text list "Banner_ManIntMsg2": 0 '**Local Message Display**'; 1 '~Spare MB2[0].1'; 2 '~Spare MB2[0].2'; 3 '~Spare MB2[0].3'; 4 '~Spare MB2[0].4'; 5 '~Spare MB2[0].5'; 6 '~Spare MB2[0].6'; 7 '~Spare MB2[0].7'; 8 '~Spare MB2[0].8'; 9 '~Spare MB2[0].9'; 10 '~Spare MB2[0].10'; 11 '~Spare MB2[0].11'; 12 '~Spare MB2[0].12'; 13 '~Spare MB2[0].13'; 14 '~Spare MB2[0].14'; 15 '~Spare MB2[0].15'; 16 '~Spare MB2[0].16'; 17 '~Spare MB2[0].17'; 18 '~Spare MB2[0].18'; 19 '~Spare MB2[0].19'; 20 '~Spare MB2[0].20'; 21 '~Spare MB2[0].21'; 22 '~Spare MB2[0].22'; 23 '~Spare MB2[0].23'; 24 '~Spare MB2[0].24'; 25 '~Spare MB2[0].25'; 26 '~Spare MB2[0].26'; 27 '~Spare MB2[0].27'; 28 '~Spare MB2[0].28'; 29 '~Spare MB2[0].29'; 30 '~Spare MB2[0].30'; 31 '~Spare MB2[0].31'; 32 '~PDPES1 - PDP EtherNet Switch Connection Inhibited MB2[1].0'; 33 '~Spare MB2[1].1'; 34 '~Spare MB2[1].2'; 35 '~MPES1 - Main Panel EtherNet Switch Connection Inhibited MB2[1].3'; 36 '~Spare MB2[1].4'; 37 '~Spare MB2[1].5'; 38 '~MPES2 - Main Panel EtherNet Switch Connection Inhibited MB2[1].6'; 39 '~Spare MB2[1].7'; 40 '~Spare MB2[1].8'; 41 '~MPES3 - Main Panel EtherNet Switch Connection Inhibited MB2[1].9'; 42 '~Spare MB2[1].10'; 43 '~Spare MB2[1].11'; 44 '~Spare MB2[1].12'; 45 '~Spare MB2[1].13'; 46 '~Spare MB2[1].14'; 47 '~Spare MB2[1].15'; 48 '~Spare MB2[1].16'; 49 '~MPES1 - Main Panel Control Power Disconnect Not On MB2[1].17'; 50 '~PDP 1 - Panel Output Disconnect Safety Switch Not On MB2[1].18'; 51 '~PDP 2 - Panel Output Disconnect Safety Switch Not On MB2[1].19'; 52 '~PDP 3 - Panel Output Disconnect Safety Switch Not On MB2[1].20'; 53 '~Spare MB2[1].21'; 54 '~Spare MB2[1].22'; 55 '~Spare MB2[1].23'; 56 '~Spare MB2[1].24'; 57 '~Spare MB2[1].25'; 58 '~Spare MB2[1].26'; 59 '~Spare MB2[1].27'; 60 '~Spare MB2[1].28'; 61 '~Spare MB2[1].29'; 62 '~Spare MB2[1].30'; 63 '~Spare MB2[1].31'; 64 '~ES3ES1 - ES3 EtherNet Switch Connection Inhibited MB2[2].0'; 65 '~Spare MB2[2].1'; 66 '~Spare MB2[2].2'; 67 '~Spare MB2[2].3'; 68 '~Spare MB2[2].4'; 69 '~Spare MB2[2].5'; 70 '~Spare MB2[2].6'; 71 '~Spare MB2[2].7'; 72 '~Spare MB2[2].8'; 73 '~ES3Sfty - Motion Control Enable Relay #1 MECR1 Still On MB2[2].9'; 74 '~ES3Sfty - Motion Control Enable Relay #1 MECR1 Not On MB2[2].10'; 75 '~ES3Sfty - Motion Control Enable Relay #2 MECR2 Still On MB2[2].11'; 76 '~ES3Sfty - Motion Control Enable Relay #2 MECR2 Not On MB2[2].12'; 77 '~ES3Sfty - EtherNet Switch Sfty Relays RESSR1 RESSR2 Not On MB2[2].13'; 78 '~ES3Sfty - EtherNet Switch Sfty Relays RESSR1 RESSR2 Still On MB2[2].14'; 79 '~Spare MB2[2].15'; 80 '~Spare MB2[2].16'; 81 '~Spare MB2[2].17'; 82 '~Spare MB2[2].18'; 83 '~Spare MB2[2].19'; 84 '~ES3 S003 Safety Gate #1 Open MB2[2].20'; 85 '~ES3 S003 Safety Gate #2 Open MB2[2].21'; 86 '~Spare MB2[2].22'; 87 '~Spare MB2[2].23'; 88 '~Spare MB2[2].24'; 89 '~Spare MB2[2].25'; 90 '~Spare MB2[2].26'; 91 '~Spare MB2[2].27'; 92 '~Spare MB2[2].28'; 93 '~Spare MB2[2].29'; 94 '~Spare MB2[2].30'; 95 '~Spare MB2[2].31'; 96 '~ES4ES1 - ES4 EtherNet Switch Connection Inhibited MB2[3].0'; 97 '~Spare MB2[3].1'; 98 '~Spare MB2[3].2'; 99 '~Spare MB2[3].3'; 100 '~Spare MB2[3].4'; 101 '~Spare MB2[3].5'; 102 '~Spare MB2[3].6'; 103 '~Spare MB2[3].7'; 104 '~Spare MB2[3].8'; 105 '~ES2Sfty - Motion Control Enable Relay #1 MECR1 Still On MB2[3].9'; 106 '~ES2Sfty - Motion Control Enable Relay #1 MECR1 Not On MB2[3].10'; 107 '~ES2Sfty - Motion Control Enable Relay #2 MECR2 Still On MB2[3].11'; 108 '~ES2Sfty - Motion Control Enable Relay #2 MECR2 Not On MB2[3].12'; 109 '~ES2Sfty - EtherNet Switch Sfty Relays RESSR1 RESSR2 Not On MB2[3].13'; 110 '~ES2Sfty - EtherNet Switch Sfty Relays RESSR1 RESSR2 Still On MB2[3].14'; 111 '~Spare MB2[3].15'; 112 '~Spare MB2[3].16'; 113 '~Spare MB2[3].17'; 114 '~Spare MB2[3].18'; 115 '~Spare MB2[3].19'; 116 '~ES2 S002 Safety Gate #1 Open MB2[3].20'; 117 '~ES2 S002 Safety Gate #2 Open MB2[3].21'; 118 '~Spare MB2[3].22'; 119 '~Spare MB2[3].23'; 120 '~Spare MB2[3].24'; 121 '~Spare MB2[3].25'; 122 '~Spare MB2[3].26'; 123 '~Spare MB2[3].27'; 124 '~Spare MB2[3].28'; 125 '~Spare MB2[3].29'; 126 '~Spare MB2[3].30'; 127 '~Spare MB2[3].31'; 128 '~PV3ES1 - PV3 EtherNet Switch Connection Inhibited MB2[4].0'; 129 '~Spare MB2[4].1'; 130 '~Spare MB2[4].2'; 131 '~Spare MB2[4].3'; 132 '~Spare MB2[4].4'; 133 '~Spare MB2[4].5'; 134 '~Spare MB2[4].6'; 135 '~Spare MB2[4].7'; 136 '~Spare MB2[4].8'; 137 '~Spare MB2[4].9'; 138 '~Spare MB2[4].10'; 139 '~PV1Sfty - EtherNet Switch Sfty Relays RESSR1 RESSR2 Not On MB2[4].11'; 140 '~PV1Sfty - EtherNet Switch Sfty Relays RESSR1 RESSR2 Still On MB2[4].12'; 141 '~Spare MB2[4].13'; 142 '~Spare MB2[4].14'; 143 '~PV1 S002 E-Stop Depressed MB2[4].15'; 144 '~PV1 S002 Safety Gate #1 Open MB2[4].16'; 145 '~PV1 S002 Safety Gate #2 Open MB2[4].17'; 146 '~Spare MB2[4].18'; 147 '~Spare MB2[4].19'; 148 '~Spare MB2[4].20'; 149 '~Spare MB2[4].21'; 150 '~Spare MB2[4].22'; 151 '~Spare MB2[4].23'; 152 '~S002 Both PanelViews Have Manual Selected MB2[4].24'; 153 '~S002 PanelView 1 Manual Selected MB2[4].25'; 154 '~Spare MB2[4].26'; 155 '~Spare MB2[4].27'; 156 '~PV1 S002 Auto Not Selected MB2[4].28'; 157 '~PV1 S002 Not In Auto Or Manual MB2[4].29'; 158 '~Spare MB2[4].30'; 159 '~Spare MB2[4].31'; 160 '~PV4ES1 - PV4 EtherNet Switch Connection Inhibited MB2[5].0'; 161 '~Spare MB2[5].1'; 162 '~Spare MB2[5].2'; 163 '~Spare MB2[5].3'; 164 '~Spare MB2[5].4'; 165 '~Spare MB2[5].5'; 166 '~Spare MB2[5].6'; 167 '~Spare MB2[5].7'; 168 '~Spare MB2[5].8'; 169 '~Spare MB2[5].9'; 170 '~Spare MB2[5].10'; 171 '~PV2Sfty - EtherNet Switch Sfty Relays RESSR1 RESSR2 Not On MB2[5].11'; 172 '~PV2Sfty - EtherNet Switch Sfty Relays RESSR1 RESSR2 Still On MB2[5].12'; 173 '~Spare MB2[5].13'; 174 '~Spare MB2[5].14'; 175 '~PV2 S002 PanelView E-Stop Depressed MB2[5].15'; 176 '~PV2 S002 Safety Gate #1 Open MB2[5].16'; 177 '~PV2 S002 Safety Gate #2 Open MB2[5].17'; 178 '~Spare MB2[5].18'; 179 '~Spare MB2[5].19'; 180 '~Spare MB2[5].20'; 181 '~Spare MB2[5].21'; 182 '~Spare MB2[5].22'; 183 '~Spare MB2[5].23'; 184 '~Spare MB2[5].24'; 185 '~S002 PanelView 2 Manual Selected MB2[5].25'; 186 '~Spare MB2[5].26'; 187 '~Spare MB2[5].27'; 188 '~PV2 S002 Auto Not Selected MB2[5].28'; 189 '~PV2 S002 Not In Auto Or Manual MB2[5].29'; 190 '~Spare MB2[5].30'; 191 '~Spare MB2[5].31'; 192 '~S001R09ES1 - S001R09 EtherNet Switch Connection Inhibited MB2[6].0'; 193 '~Spare MB2[6].1'; 194 '~Spare MB2[6].2'; 195 '~Spare MB2[6].3'; 196 '~Spare MB2[6].4'; 197 '~Spare MB2[6].5'; 198 '~Spare MB2[6].6'; 199 '~Spare MB2[6].7'; 200 '~Spare MB2[6].8'; 201 '~Spare MB2[6].9'; 202 '~Spare MB2[6].10'; 203 '~Spare MB2[6].11'; 204 '~Spare MB2[6].12'; 205 '~Spare MB2[6].13'; 206 '~Spare MB2[6].14'; 207 '~Spare MB2[6].15'; 208 '~Spare MB2[6].16'; 209 '~S001R09Sfty - Robot E-Stop Depressed MB2[6].17'; 210 '~S001R09Sfty - Robot Safety Interface Not Enabled MB2[6].18'; 211 '~S001R09Sfty - Robot DCS Has Been Edited MB2[6].19'; 212 '~S001R09CN - Robot Controller Connection Inhibited MB2[6].20'; 213 '~S001R09E#B# - Robot End Effector Module Connection Inhibited MB2[6].21'; 214 '~S001R09E#B# - Robot End Effector Module Connection Inhibited MB2[6].22'; 215 '~S001R09E#B# - Robot End Effector Module Connection Inhibited MB2[6].23'; 216 '~S001R09E#B# - Robot End Effector Module Connection Inhibited MB2[6].24'; 217 '~S001R09E#B# - Robot End Effector Module Connection Inhibited MB2[6].25'; 218 '~S001R09E#B# - Robot End Effector Module Connection Inhibited MB2[6].26'; 219 '~S001R09E#B# - Robot End Effector Module Connection Inhibited MB2[6].27'; 220 '~S001R09E#B# - Robot End Effector Module Connection Inhibited MB2[6].28'; 221 '~S001R09E#B# - Robot End Effector Module Connection Inhibited MB2[6].29'; 222 '~Spare MB2[6].30'; 223 '~Spare MB2[6].31'; 224 '~Spare MB2[7].0'; 225 '~S001R09F#B# - Robot Process I/O Connection Inhibited MB2[7].1'; 226 '~S001R09F#B# - Robot Process I/O Connection Inhibited MB2[7].2'; 227 '~S001R09F#B# - Robot Process I/O Connection Inhibited MB2[7].3'; 228 '~S001R09F#B# - Robot Process I/O Connection Inhibited MB2[7].4'; 229 '~Spare MB2[7].5'; 230 '~Spare MB2[7].6'; 231 '~Spare MB2[7].7'; 232 '~Spare MB2[7].8'; 233 '~Spare MB2[7].9'; 234 '~S001R09CN.I.Safety - Chain Fault MB2[7].10'; 235 '~S001R09CN.I.AirOn - Robot Air Not On MB2[7].11'; 236 '~S001R09CN.I.RbtAuto - Robot Not in Auto MB2[7].12'; 237 '~S001R09CN.M.InTeach - Robot In Teach MB2[7].13'; 238 '~S001R09CN.I.AtMaintPos - Robot At Maintenace MB2[7].14'; 239 '~S001R09CN.I.RunEnblInterruptAck - Robot In Hold MB2[7].15'; 240 '~S001R09CN.M.MaintPosSeld - Robot Maintenance Selected MB2[7].16'; 241 '~Spare MB2[7].17'; 242 '~Spare MB2[7].18'; 243 '~Spare MB2[7].19'; 244 '~S001R09CN.I.ExtAppCommFlt - Robot Application Communication Fault MB2[7].20'; 245 '~S001R09CN.M.AbortPickupSeld - Robot Abort Pickup Selected MB2[7].21'; 246 '~S001R09CN.M.RetFmPounceSeld - Robot Return From Pounce Selected MB2[7].22'; 247 '~S001R09CN.I.StudWld1 Comm Not OK MB2[7].23'; 248 '~S001R09CN.I.StudWld2 Comm Not OK MB2[7].24'; 249 '~S001R09CN.I.WldMode - Robot In No Weld MB2[7].25'; 250 '~S001R09CN.I.PulledTipBypSS - Robot Pulled Tip Bypass Selected MB2[7].26'; 251 '~S001R09CN.I.FlowNoFlowSS - Robot In No Flow MB2[7].27'; 252 '~S001R09CN.I.RvtNoRvtSS - Robot In No Rivet MB2[7].28'; 253 '~S001R09CN.I.WldCtrlCommOk1 - Robot Weld Controller 1 Comm Not OK MB2[7].29'; 254 '~S001R09CN.I.WldModeStud - Robot In No Weld Stud MB2[7].30'; 255 '~S001R09CN.Ix.MigWldNoWld - Robot In No Weld Mig MB2[7].31'; 256 '~S001R09CN.I.StudWld1Rdy - Robot Stud Weld Controller 1 Not Ready MB2[8].0'; 257 '~S001R09CN.I.Rvt1RdyToOperate - Robot Rivet Controller 1 Not Ready MB2[8].1'; 258 '~S001R09CN.Ix.MigRdy - Robot Mig Weld Controller Not Ready MB2[8].2'; 259 '~S001R09CN.Ix.MigWldNoWld - Robot In No Weld MB2[8].3'; 260 '~Spare MB2[8].4'; 261 '~S001R09CN.I.WldCtrlCommOk2 - Robot Weld Controller 2 Comm Not OK MB2[8].5'; 262 '~Spare MB2[8].6'; 263 '~Spare MB2[8].7'; 264 '~S001R09CN.I.StudWld2Rdy - Robot Stud Weld Controller 2 Not Ready MB2[8].8'; 265 '~S001R09CN.I.Rvt2RdyToOperate - Robot Rivet Controller 2 Not Ready MB2[8].9'; 266 '~S001R09CN.Ix.LaserWldOn - Robot Laser In No Cut MB2[8].10'; 267 '~S001R09CN.Ix.GlassNotPres - Robot Laser Glass Not Present MB2[8].11'; 268 '~S001R09CN.Ix.LaserHeadRdy - Robot Laser Head Not Ready MB2[8].12'; 269 '~S001R09CN.Ix.ChillerOn - Robot Laser Chiller Not On MB2[8].13'; 270 '~S001R09CN.Ix.GasOn - Robot Gas Not On MB2[8].14'; 271 '~S001R09 Power Meter Not Ready MB2[8].15'; 272 '~S001R09 No Wire Present Replace Barrel MB2[8].16'; 273 '~S001R09 Wire Feeder Fault Timer MB2[8].17'; 274 '~S001R09CN.Ix.NRFlt - Robot Nut Runner Not Ready MB2[8].18'; 275 '~Spare MB2[8].19'; 276 '~S001R09CN.M.WrongRivetAtNose - Remove Wrong Rivet At Nose MB2[8].20'; 277 '~S001R09CN.M.DisableRbtDrvs - In Rivet Zone But Riveter Not In Auto MB2[8].21'; 278 '~S001R09CN.I.Rvt1SystemInAuto - Rivet Controller 1 Not In Auto MB2[8].22'; 279 '~S001R09CN.I.Rvt2SystemInAuto - Rivet Controller 2 Not In Auto MB2[8].23'; 280 '~S001R09CN.M.RvtC1ReelCtr.DN - Reel Change Required MB2[8].24'; 281 '~S001R09CN.M.RvtC2ReelCtr.DN - Reel Change Required MB2[8].25'; 282 '~S001R09CN.M.AbortSkipRemain - SkipRemaining Aborted, Reset At Rbt Controller Is Required MB2[8].26'; 283 '~Spare MB2[8].27'; 284 '~Spare MB2[8].28'; 285 '~Spare MB2[8].29'; 286 '~Spare MB2[8].30'; 287 '~Spare MB2[8].31'; 288 '~Spare MB2[9].0'; 289 '~Spare MB2[9].1'; 290 '~Spare MB2[9].2'; 291 '~Spare MB2[9].3'; 292 '~Spare MB2[9].4'; 293 '~Spare MB2[9].5'; 294 '~Spare MB2[9].6'; 295 '~Spare MB2[9].7'; 296 '~Spare MB2[9].8'; 297 '~Spare MB2[9].9'; 298 '~Spare MB2[9].10'; 299 '~Spare MB2[9].11'; 300 '~Spare MB2[9].12'; 301 '~Spare MB2[9].13'; 302 '~Spare MB2[9].14'; 303 '~Spare MB2[9].15'; 304 '~Spare MB2[9].16'; 305 '~Spare MB2[9].17'; 306 '~Spare MB2[9].18'; 307 '~Spare MB2[9].19'; 308 '~Spare MB2[9].20'; 309 '~Spare MB2[9].21'; 310 '~Spare MB2[9].22'; 311 '~Spare MB2[9].23'; 312 '~Spare MB2[9].24'; 313 '~Spare MB2[9].25'; 314 '~Spare MB2[9].26'; 315 '~Spare MB2[9].27'; 316 '~Spare MB2[9].28'; 317 '~Spare MB2[9].29'; 318 '~Spare MB2[9].30'; 319 '~Spare MB2[9].31'; 320 '~Spare MB2[10].0'; 321 '~Spare MB2[10].1'; 322 '~Spare MB2[10].2'; 323 '~Spare MB2[10].3'; 324 '~Spare MB2[10].4'; 325 '~Spare MB2[10].5'; 326 '~Spare MB2[10].6'; 327 '~Spare MB2[10].7'; 328 '~Spare MB2[10].8'; 329 '~Spare MB2[10].9'; 330 '~Spare MB2[10].10'; 331 '~Spare MB2[10].11'; 332 '~Spare MB2[10].12'; 333 '~Spare MB2[10].13'; 334 '~Spare MB2[10].14'; 335 '~Spare MB2[10].15'; 336 '~Spare MB2[10].16'; 337 '~Spare MB2[10].17'; 338 '~Spare MB2[10].18'; 339 '~Spare MB2[10].19'; 340 '~Spare MB2[10].20'; 341 '~Spare MB2[10].21'; 342 '~Spare MB2[10].22'; 343 '~Spare MB2[10].23'; 344 '~Spare MB2[10].24'; 345 '~Spare MB2[10].25'; 346 '~Spare MB2[10].26'; 347 '~Spare MB2[10].27'; 348 '~Spare MB2[10].28'; 349 '~Spare MB2[10].29'; 350 '~Spare MB2[10].30'; 351 '~Spare MB2[10].31'; 352 '~Spare MB2[11].0'; 353 '~Spare MB2[11].1'; 354 '~Spare MB2[11].2'; 355 '~Spare MB2[11].3'; 356 '~Spare MB2[11].4'; 357 '~Spare MB2[11].5'; 358 '~Spare MB2[11].6'; 359 '~Spare MB2[11].7'; 360 '~Spare MB2[11].8'; 361 '~Spare MB2[11].9'; 362 '~Spare MB2[11].10'; 363 '~Spare MB2[11].11'; 364 '~Spare MB2[11].12'; 365 '~Spare MB2[11].13'; 366 '~Spare MB2[11].14'; 367 '~Spare MB2[11].15'; 368 '~Spare MB2[11].16'; 369 '~Spare MB2[11].17'; 370 '~Spare MB2[11].18'; 371 '~Spare MB2[11].19'; 372 '~Spare MB2[11].20'; 373 '~Spare MB2[11].21'; 374 '~Spare MB2[11].22'; 375 '~Spare MB2[11].23'; 376 '~Spare MB2[11].24'; 377 '~Spare MB2[11].25'; 378 '~Spare MB2[11].26'; 379 '~Spare MB2[11].27'; 380 '~Spare MB2[11].28'; 381 '~Spare MB2[11].29'; 382 '~Spare MB2[11].30'; 383 '~Spare MB2[11].31'; 384 '~S001R10ES1 - S001R10 EtherNet Switch Connection Inhibited MB2[12].0'; 385 '~Spare MB2[12].1'; 386 '~Spare MB2[12].2'; 387 '~Spare MB2[12].3'; 388 '~Spare MB2[12].4'; 389 '~Spare MB2[12].5'; 390 '~Spare MB2[12].6'; 391 '~Spare MB2[12].7'; 392 '~Spare MB2[12].8'; 393 '~Spare MB2[12].9'; 394 '~Spare MB2[12].10'; 395 '~Spare MB2[12].11'; 396 '~Spare MB2[12].12'; 397 '~Spare MB2[12].13'; 398 '~Spare MB2[12].14'; 399 '~Spare MB2[12].15'; 400 '~Spare MB2[12].16'; 401 '~S001R10Sfty - Robot E-Stop Depressed MB2[12].17'; 402 '~S001R10Sfty - Robot Safety Interface Not Enabled MB2[12].18'; 403 '~S001R10Sfty - Robot DCS Has Been Edited MB2[12].19'; 404 '~S001R10CN - Robot Controller Connection Inhibited MB2[12].20'; 405 '~S001R10E#B# - Robot End Effector Module Connection Inhibited MB2[12].21'; 406 '~S001R10E#B# - Robot End Effector Module Connection Inhibited MB2[12].22'; 407 '~S001R10E#B# - Robot End Effector Module Connection Inhibited MB2[12].23'; 408 '~S001R10E#B# - Robot End Effector Module Connection Inhibited MB2[12].24'; 409 '~S001R10E#B# - Robot End Effector Module Connection Inhibited MB2[12].25'; 410 '~S001R10E#B# - Robot End Effector Module Connection Inhibited MB2[12].26'; 411 '~S001R10E#B# - Robot End Effector Module Connection Inhibited MB2[12].27'; 412 '~S001R10E#B# - Robot End Effector Module Connection Inhibited MB2[12].28'; 413 '~S001R10E#B# - Robot End Effector Module Connection Inhibited MB2[12].29'; 414 '~Spare MB2[12].30'; 415 '~Spare MB2[12].31'; 416 '~Spare MB2[13].0'; 417 '~S001R10F#B# - Robot Process I/O Connection Inhibited MB2[13].1'; 418 '~S001R10F#B# - Robot Process I/O Connection Inhibited MB2[13].2'; 419 '~S001R10F#B# - Robot Process I/O Connection Inhibited MB2[13].3'; 420 '~S001R10F#B# - Robot Process I/O Connection Inhibited MB2[13].4'; 421 '~Spare MB2[13].5'; 422 '~Spare MB2[13].6'; 423 '~Spare MB2[13].7'; 424 '~Spare MB2[13].8'; 425 '~Spare MB2[13].9'; 426 '~S001R10CN.I.Safety - Chain Fault MB2[13].10'; 427 '~S001R10CN.I.AirOn - Robot Air Not On MB2[13].11'; 428 '~S001R10CN.I.RbtAuto - Robot Not in Auto MB2[13].12'; 429 '~S001R10CN.M.InTeach - Robot In Teach MB2[13].13'; 430 '~S001R10CN.I.AtMaintPos - Robot At Maintenace MB2[13].14'; 431 '~S001R10CN.I.RunEnblInterruptAck - Robot In Hold MB2[13].15'; 432 '~S001R10CN.M.MaintPosSeld - Robot Maintenance Selected MB2[13].16'; 433 '~Spare MB2[13].17'; 434 '~Spare MB2[13].18'; 435 '~Spare MB2[13].19'; 436 '~S001R10CN.I.ExtAppCommFlt - Robot Application Communication Fault MB2[13].20'; 437 '~S001R10CN.M.AbortPickupSeld - Robot Abort Pickup Selected MB2[13].21'; 438 '~S001R10CN.M.RetFmPounceSeld - Robot Return From Pounce Selected MB2[13].22'; 439 '~S001R10CN.I.StudWld1 Comm Not OK MB2[13].23'; 440 '~S001R10CN.I.StudWld2 Comm Not OK MB2[13].24'; 441 '~S001R10CN.I.WldMode - Robot In No Weld MB2[13].25'; 442 '~S001R10CN.I.PulledTipBypSS - Robot Pulled Tip Bypass Selected MB2[13].26'; 443 '~S001R10CN.I.FlowNoFlowSS - Robot In No Flow MB2[13].27'; 444 '~S001R10CN.I.RvtNoRvtSS - Robot In No Rivet MB2[13].28'; 445 '~S001R10CN.I.WldCtrlCommOk1 - Robot Weld Controller 1 Comm Not OK MB2[13].29'; 446 '~S001R10CN.I.WldModeStud - Robot In No Weld Stud MB2[13].30'; 447 '~S001R10CN.Ix.MigWldNoWld - Robot In No Weld Mig MB2[13].31'; 448 '~S001R10CN.I.StudWld1Rdy - Robot Stud Weld Controller 1 Not Ready MB2[14].0'; 449 '~S001R10CN.I.Rvt1RdyToOperate - Robot Rivet Controller 1 Not Ready MB2[14].1'; 450 '~S001R10CN.Ix.MigRdy - Robot Mig Weld Controller Not Ready MB2[14].2'; 451 '~S001R10CN.Ix.MigWldNoWld - Robot In No Weld MB2[14].3'; 452 '~Spare MB2[14].4'; 453 '~S001R10CN.I.WldCtrlCommOk2 - Robot Weld Controller 2 Comm Not OK MB2[14].5'; 454 '~Spare MB2[14].6'; 455 '~Spare MB2[14].7'; 456 '~S001R10CN.I.StudWld2Rdy - Robot Stud Weld Controller 2 Not Ready MB2[14].8'; 457 '~S001R10CN.I.Rvt2RdyToOperate - Robot Rivet Controller 2 Not Ready MB2[14].9'; 458 '~S001R10CN.Ix.LaserWldOn - Robot Laser In No Cut MB2[14].10'; 459 '~S001R10CN.Ix.GlassNotPres - Robot Laser Glass Not Present MB2[14].11'; 460 '~S001R10CN.Ix.LaserHeadRdy - Robot Laser Head Not Ready MB2[14].12'; 461 '~S001R10CN.Ix.ChillerOn - Robot Laser Chiller Not On MB2[14].13'; 462 '~S001R10CN.Ix.GasOn - Robot Gas Not On MB2[14].14'; 463 '~S001R10 Power Meter Not Ready MB2[14].15'; 464 '~S001R10 No Wire Present Replace Barrel MB2[14].16'; 465 '~S001R10 Wire Feeder Fault Timer MB2[14].17'; 466 '~S001R10CN.Ix.NRFlt - Robot Nut Runner Not Ready MB2[14].18'; 467 '~Spare MB2[14].19'; 468 '~S001R10CN.M.WrongRivetAtNose - Remove Wrong Rivet At Nose MB2[14].20'; 469 '~S001R10CN.M.DisableRbtDrvs - In Rivet Zone But Riveter Not In Auto MB2[14].21'; 470 '~S001R10CN.I.Rvt1SystemInAuto - Rivet Controller 1 Not In Auto MB2[14].22'; 471 '~S001R10CN.I.Rvt2SystemInAuto - Rivet Controller 2 Not In Auto MB2[14].23'; 472 '~S001R10CN.M.RvtC1ReelCtr.DN - Reel Change Required MB2[14].24'; 473 '~S001R10CN.M.RvtC2ReelCtr.DN - Reel Change Required MB2[14].25'; 474 '~S001R10CN.M.AbortSkipRemain - SkipRemaining Aborted, Reset At Rbt Controller Is Required MB2[14].26'; 475 '~Spare MB2[14].27'; 476 '~Spare MB2[14].28'; 477 '~Spare MB2[14].29'; 478 '~Spare MB2[14].30'; 479 '~Spare MB2[14].31'; 480 '~Spare MB2[15].0'; 481 '~Spare MB2[15].1'; 482 '~Spare MB2[15].2'; 483 '~Spare MB2[15].3'; 484 '~Spare MB2[15].4'; 485 '~Spare MB2[15].5'; 486 '~Spare MB2[15].6'; 487 '~Spare MB2[15].7'; 488 '~Spare MB2[15].8'; 489 '~Spare MB2[15].9'; 490 '~Spare MB2[15].10'; 491 '~Spare MB2[15].11'; 492 '~Spare MB2[15].12'; 493 '~Spare MB2[15].13'; 494 '~Spare MB2[15].14'; 495 '~Spare MB2[15].15'; 496 '~Spare MB2[15].16'; 497 '~Spare MB2[15].17'; 498 '~Spare MB2[15].18'; 499 '~Spare MB2[15].19'; 500 '~Spare MB2[15].20'; 501 '~Spare MB2[15].21'; 502 '~Spare MB2[15].22'; 503 '~Spare MB2[15].23'; 504 '~Spare MB2[15].24'; 505 '~Spare MB2[15].25'; 506 '~Spare MB2[15].26'; 507 '~Spare MB2[15].27'; 508 '~Spare MB2[15].28'; 509 '~Spare MB2[15].29'; 510 '~Spare MB2[15].30'; 511 '~Spare MB2[15].31'; 512 '~Spare MB2[16].0'; 513 '~Spare MB2[16].1'; 514 '~Spare MB2[16].2'; 515 '~Spare MB2[16].3'; 516 '~Spare MB2[16].4'; 517 '~Spare MB2[16].5'; 518 '~Spare MB2[16].6'; 519 '~Spare MB2[16].7'; 520 '~Spare MB2[16].8'; 521 '~Spare MB2[16].9'; 522 '~Spare MB2[16].10'; 523 '~Spare MB2[16].11'; 524 '~Spare MB2[16].12'; 525 '~Spare MB2[16].13'; 526 '~Spare MB2[16].14'; 527 '~Spare MB2[16].15'; 528 '~Spare MB2[16].16'; 529 '~Spare MB2[16].17'; 530 '~Spare MB2[16].18'; 531 '~Spare MB2[16].19'; 532 '~Spare MB2[16].20'; 533 '~Spare MB2[16].21'; 534 '~Spare MB2[16].22'; 535 '~Spare MB2[16].23'; 536 '~Spare MB2[16].24'; 537 '~Spare MB2[16].25'; 538 '~Spare MB2[16].26'; 539 '~Spare MB2[16].27'; 540 '~Spare MB2[16].28'; 541 '~Spare MB2[16].29'; 542 '~Spare MB2[16].30'; 543 '~Spare MB2[16].31'; 544 '~Spare MB2[17].0'; 545 '~Spare MB2[17].1'; 546 '~Spare MB2[17].2'; 547 '~Spare MB2[17].3'; 548 '~Spare MB2[17].4'; 549 '~Spare MB2[17].5'; 550 '~Spare MB2[17].6'; 551 '~Spare MB2[17].7'; 552 '~Spare MB2[17].8'; 553 '~Spare MB2[17].9'; 554 '~Spare MB2[17].10'; 555 '~Spare MB2[17].11'; 556 '~Spare MB2[17].12'; 557 '~Spare MB2[17].13'; 558 '~Spare MB2[17].14'; 559 '~Spare MB2[17].15'; 560 '~Spare MB2[17].16'; 561 '~Spare MB2[17].17'; 562 '~Spare MB2[17].18'; 563 '~Spare MB2[17].19'; 564 '~Spare MB2[17].20'; 565 '~Spare MB2[17].21'; 566 '~Spare MB2[17].22'; 567 '~Spare MB2[17].23'; 568 '~Spare MB2[17].24'; 569 '~Spare MB2[17].25'; 570 '~Spare MB2[17].26'; 571 '~Spare MB2[17].27'; 572 '~Spare MB2[17].28'; 573 '~Spare MB2[17].29'; 574 '~Spare MB2[17].30'; 575 '~Spare MB2[17].31'; 576 '~S001R11ES1 - S001R11 EtherNet Switch Connection Inhibited MB2[18].0'; 577 '~Spare MB2[18].1'; 578 '~Spare MB2[18].2'; 579 '~Spare MB2[18].3'; 580 '~Spare MB2[18].4'; 581 '~Spare MB2[18].5'; 582 '~Spare MB2[18].6'; 583 '~Spare MB2[18].7'; 584 '~Spare MB2[18].8'; 585 '~Spare MB2[18].9'; 586 '~Spare MB2[18].10'; 587 '~Spare MB2[18].11'; 588 '~Spare MB2[18].12'; 589 '~Spare MB2[18].13'; 590 '~Spare MB2[18].14'; 591 '~Spare MB2[18].15'; 592 '~Spare MB2[18].16'; 593 '~S001R11Sfty - Robot E-Stop Depressed MB2[18].17'; 594 '~S001R11Sfty - Robot Safety Interface Not Enabled MB2[18].18'; 595 '~S001R11Sfty - Robot DCS Has Been Edited MB2[18].19'; 596 '~S001R11CN - Robot Controller Connection Inhibited MB2[18].20'; 597 '~S001R11E#B# - Robot End Effector Module Connection Inhibited MB2[18].21'; 598 '~S001R11E#B# - Robot End Effector Module Connection Inhibited MB2[18].22'; 599 '~S001R11E#B# - Robot End Effector Module Connection Inhibited MB2[18].23'; 600 '~S001R11E#B# - Robot End Effector Module Connection Inhibited MB2[18].24'; 601 '~S001R11E#B# - Robot End Effector Module Connection Inhibited MB2[18].25'; 602 '~S001R11E#B# - Robot End Effector Module Connection Inhibited MB2[18].26'; 603 '~S001R11E#B# - Robot End Effector Module Connection Inhibited MB2[18].27'; 604 '~S001R11E#B# - Robot End Effector Module Connection Inhibited MB2[18].28'; 605 '~S001R11E#B# - Robot End Effector Module Connection Inhibited MB2[18].29'; 606 '~Spare MB2[18].30'; 607 '~Spare MB2[18].31'; 608 '~Spare MB2[19].0'; 609 '~S001R11F#B# - Robot Process I/O Connection Inhibited MB2[19].1'; 610 '~S001R11F#B# - Robot Process I/O Connection Inhibited MB2[19].2'; 611 '~S001R11F#B# - Robot Process I/O Connection Inhibited MB2[19].3'; 612 '~S001R11F#B# - Robot Process I/O Connection Inhibited MB2[19].4'; 613 '~Spare MB2[19].5'; 614 '~Spare MB2[19].6'; 615 '~Spare MB2[19].7'; 616 '~Spare MB2[19].8'; 617 '~Spare MB2[19].9'; 618 '~S001R11CN.I.Safety - Chain Fault MB2[19].10'; 619 '~S001R11CN.I.AirOn - Robot Air Not On MB2[19].11'; 620 '~S001R11CN.I.RbtAuto - Robot Not in Auto MB2[19].12'; 621 '~S001R11CN.M.InTeach - Robot In Teach MB2[19].13'; 622 '~S001R11CN.I.AtMaintPos - Robot At Maintenace MB2[19].14'; 623 '~S001R11CN.I.RunEnblInterruptAck - Robot In Hold MB2[19].15'; 624 '~S001R11CN.M.MaintPosSeld - Robot Maintenance Selected MB2[19].16'; 625 '~Spare MB2[19].17'; 626 '~Spare MB2[19].18'; 627 '~Spare MB2[19].19'; 628 '~S001R11CN.I.ExtAppCommFlt - Robot Application Communication Fault MB2[19].20'; 629 '~S001R11CN.M.AbortPickupSeld - Robot Abort Pickup Selected MB2[19].21'; 630 '~S001R11CN.M.RetFmPounceSeld - Robot Return From Pounce Selected MB2[19].22'; 631 '~S001R11CN.I.StudWld1 Comm Not OK MB2[19].23'; 632 '~S001R11CN.I.StudWld2 Comm Not OK MB2[19].24'; 633 '~S001R11CN.I.WldMode - Robot In No Weld MB2[19].25'; 634 '~S001R11CN.I.PulledTipBypSS - Robot Pulled Tip Bypass Selected MB2[19].26'; 635 '~S001R11CN.I.FlowNoFlowSS - Robot In No Flow MB2[19].27'; 636 '~S001R11CN.I.RvtNoRvtSS - Robot In No Rivet MB2[19].28'; 637 '~S001R11CN.I.WldCtrlCommOk1 - Robot Weld Controller 1 Comm Not OK MB2[19].29'; 638 '~S001R11CN.I.WldModeStud - Robot In No Weld Stud MB2[19].30'; 639 '~S001R11CN.Ix.MigWldNoWld - Robot In No Weld Mig MB2[19].31'; 640 '~S001R11CN.I.StudWld1Rdy - Robot Stud Weld Controller 1 Not Ready MB2[20].0'; 641 '~S001R11CN.I.Rvt1RdyToOperate - Robot Rivet Controller 1 Not Ready MB2[20].1'; 642 '~S001R11CN.Ix.MigRdy - Robot Mig Weld Controller Not Ready MB2[20].2'; 643 '~S001R11CN.Ix.MigWldNoWld - Robot In No Weld MB2[20].3'; 644 '~Spare MB2[20].4'; 645 '~S001R11CN.I.WldCtrlCommOk2 - Robot Weld Controller 2 Comm Not OK MB2[20].5'; 646 '~Spare MB2[20].6'; 647 '~Spare MB2[20].7'; 648 '~S001R11CN.I.StudWld2Rdy - Robot Stud Weld Controller 2 Not Ready MB2[20].8'; 649 '~S001R11CN.I.Rvt2RdyToOperate - Robot Rivet Controller 2 Not Ready MB2[20].9'; 650 '~S001R11CN.Ix.LaserWldOn - Robot Laser In No Cut MB2[20].10'; 651 '~S001R11CN.Ix.GlassNotPres - Robot Laser Glass Not Present MB2[20].11'; 652 '~S001R11CN.Ix.LaserHeadRdy - Robot Laser Head Not Ready MB2[20].12'; 653 '~S001R11CN.Ix.ChillerOn - Robot Laser Chiller Not On MB2[20].13'; 654 '~S001R11CN.Ix.GasOn - Robot Gas Not On MB2[20].14'; 655 '~S001R11 Power Meter Not Ready MB2[20].15'; 656 '~S001R11 No Wire Present Replace Barrel MB2[20].16'; 657 '~S001R11 Wire Feeder Fault Timer MB2[20].17'; 658 '~S001R11CN.Ix.NRFlt - Robot Nut Runner Not Ready MB2[20].18'; 659 '~Spare MB2[20].19'; 660 '~S001R11CN.M.WrongRivetAtNose - Remove Wrong Rivet At Nose MB2[20].20'; 661 '~S001R11CN.M.DisableRbtDrvs - In Rivet Zone But Riveter Not In Auto MB2[20].21'; 662 '~S001R11CN.I.Rvt1SystemInAuto - Rivet Controller 1 Not In Auto MB2[20].22'; 663 '~S001R11CN.I.Rvt2SystemInAuto - Rivet Controller 2 Not In Auto MB2[20].23'; 664 '~S001R11CN.M.RvtC1ReelCtr.DN - Reel Change Required MB2[20].24'; 665 '~S001R11CN.M.RvtC2ReelCtr.DN - Reel Change Required MB2[20].25'; 666 '~S001R11CN.M.AbortSkipRemain - SkipRemaining Aborted, Reset At Rbt Controller Is Required MB2[20].26'; 667 '~Spare MB2[20].27'; 668 '~Spare MB2[20].28'; 669 '~Spare MB2[20].29'; 670 '~Spare MB2[20].30'; 671 '~Spare MB2[20].31'; 672 '~Spare MB2[21].0'; 673 '~Spare MB2[21].1'; 674 '~Spare MB2[21].2'; 675 '~Spare MB2[21].3'; 676 '~Spare MB2[21].4'; 677 '~Spare MB2[21].5'; 678 '~Spare MB2[21].6'; 679 '~Spare MB2[21].7'; 680 '~Spare MB2[21].8'; 681 '~Spare MB2[21].9'; 682 '~Spare MB2[21].10'; 683 '~Spare MB2[21].11'; 684 '~Spare MB2[21].12'; 685 '~Spare MB2[21].13'; 686 '~Spare MB2[21].14'; 687 '~Spare MB2[21].15'; 688 '~Spare MB2[21].16'; 689 '~Spare MB2[21].17'; 690 '~Spare MB2[21].18'; 691 '~Spare MB2[21].19'; 692 '~Spare MB2[21].20'; 693 '~Spare MB2[21].21'; 694 '~Spare MB2[21].22'; 695 '~Spare MB2[21].23'; 696 '~Spare MB2[21].24'; 697 '~Spare MB2[21].25'; 698 '~Spare MB2[21].26'; 699 '~Spare MB2[21].27'; 700 '~Spare MB2[21].28'; 701 '~Spare MB2[21].29'; 702 '~Spare MB2[21].30'; 703 '~Spare MB2[21].31'; 704 '~Spare MB2[22].0'; 705 '~Spare MB2[22].1'; 706 '~Spare MB2[22].2'; 707 '~Spare MB2[22].3'; 708 '~Spare MB2[22].4'; 709 '~Spare MB2[22].5'; 710 '~Spare MB2[22].6'; 711 '~Spare MB2[22].7'; 712 '~Spare MB2[22].8'; 713 '~Spare MB2[22].9'; 714 '~Spare MB2[22].10'; 715 '~Spare MB2[22].11'; 716 '~Spare MB2[22].12'; 717 '~Spare MB2[22].13'; 718 '~Spare MB2[22].14'; 719 '~Spare MB2[22].15'; 720 '~Spare MB2[22].16'; 721 '~Spare MB2[22].17'; 722 '~Spare MB2[22].18'; 723 '~Spare MB2[22].19'; 724 '~Spare MB2[22].20'; 725 '~Spare MB2[22].21'; 726 '~Spare MB2[22].22'; 727 '~Spare MB2[22].23'; 728 '~Spare MB2[22].24'; 729 '~Spare MB2[22].25'; 730 '~Spare MB2[22].26'; 731 '~Spare MB2[22].27'; 732 '~Spare MB2[22].28'; 733 '~Spare MB2[22].29'; 734 '~Spare MB2[22].30'; 735 '~Spare MB2[22].31'; 736 '~Spare MB2[23].0'; 737 '~Spare MB2[23].1'; 738 '~Spare MB2[23].2'; 739 '~Spare MB2[23].3'; 740 '~Spare MB2[23].4'; 741 '~Spare MB2[23].5'; 742 '~Spare MB2[23].6'; 743 '~Spare MB2[23].7'; 744 '~Spare MB2[23].8'; 745 '~Spare MB2[23].9'; 746 '~Spare MB2[23].10'; 747 '~Spare MB2[23].11'; 748 '~Spare MB2[23].12'; 749 '~Spare MB2[23].13'; 750 '~Spare MB2[23].14'; 751 '~Spare MB2[23].15'; 752 '~Spare MB2[23].16'; 753 '~Spare MB2[23].17'; 754 '~Spare MB2[23].18'; 755 '~Spare MB2[23].19'; 756 '~Spare MB2[23].20'; 757 '~Spare MB2[23].21'; 758 '~Spare MB2[23].22'; 759 '~Spare MB2[23].23'; 760 '~Spare MB2[23].24'; 761 '~Spare MB2[23].25'; 762 '~Spare MB2[23].26'; 763 '~Spare MB2[23].27'; 764 '~Spare MB2[23].28'; 765 '~Spare MB2[23].29'; 766 '~Spare MB2[23].30'; 767 '~Spare MB2[23].31'; 768 '~S001R12ES1 - S001R12 EtherNet Switch Connection Inhibited MB2[24].0'; 769 '~Spare MB2[24].1'; 770 '~Spare MB2[24].2'; 771 '~Spare MB2[24].3'; 772 '~Spare MB2[24].4'; 773 '~Spare MB2[24].5'; 774 '~Spare MB2[24].6'; 775 '~Spare MB2[24].7'; 776 '~Spare MB2[24].8'; 777 '~Spare MB2[24].9'; 778 '~Spare MB2[24].10'; 779 '~Spare MB2[24].11'; 780 '~Spare MB2[24].12'; 781 '~Spare MB2[24].13'; 782 '~Spare MB2[24].14'; 783 '~Spare MB2[24].15'; 784 '~Spare MB2[24].16'; 785 '~S001R12Sfty - Robot E-Stop Depressed MB2[24].17'; 786 '~S001R12Sfty - Robot Safety Interface Not Enabled MB2[24].18'; 787 '~S001R12Sfty - Robot DCS Has Been Edited MB2[24].19'; 788 '~S001R12CN - Robot Controller Connection Inhibited MB2[24].20'; 789 '~S001R12E#B# - Robot End Effector Module Connection Inhibited MB2[24].21'; 790 '~S001R12E#B# - Robot End Effector Module Connection Inhibited MB2[24].22'; 791 '~S001R12E#B# - Robot End Effector Module Connection Inhibited MB2[24].23'; 792 '~S001R12E#B# - Robot End Effector Module Connection Inhibited MB2[24].24'; 793 '~S001R12E#B# - Robot End Effector Module Connection Inhibited MB2[24].25'; 794 '~S001R12E#B# - Robot End Effector Module Connection Inhibited MB2[24].26'; 795 '~S001R12E#B# - Robot End Effector Module Connection Inhibited MB2[24].27'; 796 '~S001R12E#B# - Robot End Effector Module Connection Inhibited MB2[24].28'; 797 '~S001R12E#B# - Robot End Effector Module Connection Inhibited MB2[24].29'; 798 '~Spare MB2[24].30'; 799 '~Spare MB2[24].31'; 800 '~Spare MB2[25].0'; 801 '~S001R12F#B# - Robot Process I/O Connection Inhibited MB2[25].1'; 802 '~S001R12F#B# - Robot Process I/O Connection Inhibited MB2[25].2'; 803 '~S001R12F#B# - Robot Process I/O Connection Inhibited MB2[25].3'; 804 '~S001R12F#B# - Robot Process I/O Connection Inhibited MB2[25].4'; 805 '~Spare MB2[25].5'; 806 '~Spare MB2[25].6'; 807 '~Spare MB2[25].7'; 808 '~Spare MB2[25].8'; 809 '~Spare MB2[25].9'; 810 '~S001R12CN.I.Safety - Chain Fault MB2[25].10'; 811 '~S001R12CN.I.AirOn - Robot Air Not On MB2[25].11'; 812 '~S001R12CN.I.RbtAuto - Robot Not in Auto MB2[25].12'; 813 '~S001R12CN.M.InTeach - Robot In Teach MB2[25].13'; 814 '~S001R12CN.I.AtMaintPos - Robot At Maintenace MB2[25].14'; 815 '~S001R12CN.I.RunEnblInterruptAck - Robot In Hold MB2[25].15'; 816 '~S001R12CN.M.MaintPosSeld - Robot Maintenance Selected MB2[25].16'; 817 '~Spare MB2[25].17'; 818 '~Spare MB2[25].18'; 819 '~Spare MB2[25].19'; 820 '~S001R12CN.I.ExtAppCommFlt - Robot Application Communication Fault MB2[25].20'; 821 '~S001R12CN.M.AbortPickupSeld - Robot Abort Pickup Selected MB2[25].21'; 822 '~S001R12CN.M.RetFmPounceSeld - Robot Return From Pounce Selected MB2[25].22'; 823 '~S001R12CN.I.StudWld1 Comm Not OK MB2[25].23'; 824 '~S001R12CN.I.StudWld2 Comm Not OK MB2[25].24'; 825 '~S001R12CN.I.WldMode - Robot In No Weld MB2[25].25'; 826 '~S001R12CN.I.PulledTipBypSS - Robot Pulled Tip Bypass Selected MB2[25].26'; 827 '~S001R12CN.I.FlowNoFlowSS - Robot In No Flow MB2[25].27'; 828 '~S001R12CN.I.RvtNoRvtSS - Robot In No Rivet MB2[25].28'; 829 '~S001R12CN.I.WldCtrlCommOk1 - Robot Weld Controller 1 Comm Not OK MB2[25].29'; 830 '~S001R12CN.I.WldModeStud - Robot In No Weld Stud MB2[25].30'; 831 '~S001R12CN.Ix.MigWldNoWld - Robot In No Weld Mig MB2[25].31'; 832 '~S001R12CN.I.StudWld1Rdy - Robot Stud Weld Controller 1 Not Ready MB2[26].0'; 833 '~S001R12CN.I.Rvt1RdyToOperate - Robot Rivet Controller 1 Not Ready MB2[26].1'; 834 '~S001R12CN.Ix.MigRdy - Robot Mig Weld Controller Not Ready MB2[26].2'; 835 '~S001R12CN.Ix.MigWldNoWld - Robot In No Weld MB2[26].3'; 836 '~Spare MB2[26].4'; 837 '~S001R12CN.I.WldCtrlCommOk2 - Robot Weld Controller 2 Comm Not OK MB2[26].5'; 838 '~Spare MB2[26].6'; 839 '~Spare MB2[26].7'; 840 '~S001R12CN.I.StudWld2Rdy - Robot Stud Weld Controller 2 Not Ready MB2[26].8'; 841 '~S001R12CN.I.Rvt2RdyToOperate - Robot Rivet Controller 2 Not Ready MB2[26].9'; 842 '~S001R12CN.Ix.LaserWldOn - Robot Laser In No Cut MB2[26].10'; 843 '~S001R12CN.Ix.GlassNotPres - Robot Laser Glass Not Present MB2[26].11'; 844 '~S001R12CN.Ix.LaserHeadRdy - Robot Laser Head Not Ready MB2[26].12'; 845 '~S001R12CN.Ix.ChillerOn - Robot Laser Chiller Not On MB2[26].13'; 846 '~S001R12CN.Ix.GasOn - Robot Gas Not On MB2[26].14'; 847 '~S001R12 Power Meter Not Ready MB2[26].15'; 848 '~S001R12 No Wire Present Replace Barrel MB2[26].16'; 849 '~S001R12 Wire Feeder Fault Timer MB2[26].17'; 850 '~S001R12CN.Ix.NRFlt - Robot Nut Runner Not Ready MB2[26].18'; 851 '~Spare MB2[26].19'; 852 '~S001R12CN.M.WrongRivetAtNose - Remove Wrong Rivet At Nose MB2[26].20'; 853 '~S001R12CN.M.DisableRbtDrvs - In Rivet Zone But Riveter Not In Auto MB2[26].21'; 854 '~S001R12CN.I.Rvt1SystemInAuto - Rivet Controller 1 Not In Auto MB2[26].22'; 855 '~S001R12CN.I.Rvt2SystemInAuto - Rivet Controller 2 Not In Auto MB2[26].23'; 856 '~S001R12CN.M.RvtC1ReelCtr.DN - Reel Change Required MB2[26].24'; 857 '~S001R12CN.M.RvtC2ReelCtr.DN - Reel Change Required MB2[26].25'; 858 '~S001R12CN.M.AbortSkipRemain - SkipRemaining Aborted, Reset At Rbt Controller Is Required MB2[26].26'; 859 '~Spare MB2[26].27'; 860 '~Spare MB2[26].28'; 861 '~Spare MB2[26].29'; 862 '~Spare MB2[26].30'; 863 '~Spare MB2[26].31'; 864 '~Spare MB2[27].0'; 865 '~Spare MB2[27].1'; 866 '~Spare MB2[27].2'; 867 '~Spare MB2[27].3'; 868 '~Spare MB2[27].4'; 869 '~Spare MB2[27].5'; 870 '~Spare MB2[27].6'; 871 '~Spare MB2[27].7'; 872 '~Spare MB2[27].8'; 873 '~Spare MB2[27].9'; 874 '~Spare MB2[27].10'; 875 '~Spare MB2[27].11'; 876 '~Spare MB2[27].12'; 877 '~Spare MB2[27].13'; 878 '~Spare MB2[27].14'; 879 '~Spare MB2[27].15'; 880 '~Spare MB2[27].16'; 881 '~Spare MB2[27].17'; 882 '~Spare MB2[27].18'; 883 '~Spare MB2[27].19'; 884 '~Spare MB2[27].20'; 885 '~Spare MB2[27].21'; 886 '~Spare MB2[27].22'; 887 '~Spare MB2[27].23'; 888 '~Spare MB2[27].24'; 889 '~Spare MB2[27].25'; 890 '~Spare MB2[27].26'; 891 '~Spare MB2[27].27'; 892 '~Spare MB2[27].28'; 893 '~Spare MB2[27].29'; 894 '~Spare MB2[27].30'; 895 '~Spare MB2[27].31'; 896 '~Spare MB2[28].0'; 897 '~Spare MB2[28].1'; 898 '~Spare MB2[28].2'; 899 '~Spare MB2[28].3'; 900 '~Spare MB2[28].4'; 901 '~Spare MB2[28].5'; 902 '~Spare MB2[28].6'; 903 '~Spare MB2[28].7'; 904 '~Spare MB2[28].8'; 905 '~Spare MB2[28].9'; 906 '~Spare MB2[28].10'; 907 '~Spare MB2[28].11'; 908 '~Spare MB2[28].12'; 909 '~Spare MB2[28].13'; 910 '~Spare MB2[28].14'; 911 '~Spare MB2[28].15'; 912 '~Spare MB2[28].16'; 913 '~Spare MB2[28].17'; 914 '~Spare MB2[28].18'; 915 '~Spare MB2[28].19'; 916 '~Spare MB2[28].20'; 917 '~Spare MB2[28].21'; 918 '~Spare MB2[28].22'; 919 '~Spare MB2[28].23'; 920 '~Spare MB2[28].24'; 921 '~Spare MB2[28].25'; 922 '~Spare MB2[28].26'; 923 '~Spare MB2[28].27'; 924 '~Spare MB2[28].28'; 925 '~Spare MB2[28].29'; 926 '~Spare MB2[28].30'; 927 '~Spare MB2[28].31'; 928 '~Spare MB2[29].0'; 929 '~Spare MB2[29].1'; 930 '~Spare MB2[29].2'; 931 '~Spare MB2[29].3'; 932 '~Spare MB2[29].4'; 933 '~Spare MB2[29].5'; 934 '~Spare MB2[29].6'; 935 '~Spare MB2[29].7'; 936 '~Spare MB2[29].8'; 937 '~Spare MB2[29].9'; 938 '~Spare MB2[29].10'; 939 '~Spare MB2[29].11'; 940 '~Spare MB2[29].12'; 941 '~Spare MB2[29].13'; 942 '~Spare MB2[29].14'; 943 '~Spare MB2[29].15'; 944 '~Spare MB2[29].16'; 945 '~Spare MB2[29].17'; 946 '~Spare MB2[29].18'; 947 '~Spare MB2[29].19'; 948 '~Spare MB2[29].20'; 949 '~Spare MB2[29].21'; 950 '~Spare MB2[29].22'; 951 '~Spare MB2[29].23'; 952 '~Spare MB2[29].24'; 953 '~Spare MB2[29].25'; 954 '~Spare MB2[29].26'; 955 '~Spare MB2[29].27'; 956 '~Spare MB2[29].28'; 957 '~Spare MB2[29].29'; 958 '~Spare MB2[29].30'; 959 '~Spare MB2[29].31'; 960 '~S001R13ES1 - S001R13 EtherNet Switch Connection Inhibited MB2[30].0'; 961 '~Spare MB2[30].1'; 962 '~Spare MB2[30].2'; 963 '~Spare MB2[30].3'; 964 '~Spare MB2[30].4'; 965 '~Spare MB2[30].5'; 966 '~Spare MB2[30].6'; 967 '~Spare MB2[30].7'; 968 '~Spare MB2[30].8'; 969 '~Spare MB2[30].9'; 970 '~Spare MB2[30].10'; 971 '~Spare MB2[30].11'; 972 '~Spare MB2[30].12'; 973 '~Spare MB2[30].13'; 974 '~Spare MB2[30].14'; 975 '~Spare MB2[30].15'; 976 '~Spare MB2[30].16'; 977 '~S001R13Sfty - Robot E-Stop Depressed MB2[30].17'; 978 '~S001R13Sfty - Robot Safety Interface Not Enabled MB2[30].18'; 979 '~S001R13Sfty - Robot DCS Has Been Edited MB2[30].19'; 980 '~S001R13CN - Robot Controller Connection Inhibited MB2[30].20'; 981 '~S001R13E#B# - Robot End Effector Module Connection Inhibited MB2[30].21'; 982 '~S001R13E#B# - Robot End Effector Module Connection Inhibited MB2[30].22'; 983 '~S001R13E#B# - Robot End Effector Module Connection Inhibited MB2[30].23'; 984 '~S001R13E#B# - Robot End Effector Module Connection Inhibited MB2[30].24'; 985 '~S001R13E#B# - Robot End Effector Module Connection Inhibited MB2[30].25'; 986 '~S001R13E#B# - Robot End Effector Module Connection Inhibited MB2[30].26'; 987 '~S001R13E#B# - Robot End Effector Module Connection Inhibited MB2[30].27'; 988 '~S001R13E#B# - Robot End Effector Module Connection Inhibited MB2[30].28'; 989 '~S001R13E#B# - Robot End Effector Module Connection Inhibited MB2[30].29'; 990 '~Spare MB2[30].30'; 991 '~Spare MB2[30].31'; 992 '~Spare MB2[31].0'; 993 '~S001R13F#B# - Robot Process I/O Connection Inhibited MB2[31].1'; 994 '~S001R13F#B# - Robot Process I/O Connection Inhibited MB2[31].2'; 995 '~S001R13F#B# - Robot Process I/O Connection Inhibited MB2[31].3'; 996 '~S001R13F#B# - Robot Process I/O Connection Inhibited MB2[31].4'; 997 '~Spare MB2[31].5'; 998 '~Spare MB2[31].6'; 999 '~Spare MB2[31].7'; 1000 '~Spare MB2[31].8'; 1001 '~Spare MB2[31].9'; 1002 '~S001R13CN.I.Safety - Chain Fault MB2[31].10'; 1003 '~S001R13CN.I.AirOn - Robot Air Not On MB2[31].11'; 1004 '~S001R13CN.I.RbtAuto - Robot Not in Auto MB2[31].12'; 1005 '~S001R13CN.M.InTeach - Robot In Teach MB2[31].13'; 1006 '~S001R13CN.I.AtMaintPos - Robot At Maintenace MB2[31].14'; 1007 '~S001R13CN.I.RunEnblInterruptAck - Robot In Hold MB2[31].15'; 1008 '~S001R13CN.M.MaintPosSeld - Robot Maintenance Selected MB2[31].16'; 1009 '~Spare MB2[31].17'; 1010 '~Spare MB2[31].18'; 1011 '~Spare MB2[31].19'; 1012 '~S001R13CN.I.ExtAppCommFlt - Robot Application Communication Fault MB2[31].20'; 1013 '~S001R13CN.M.AbortPickupSeld - Robot Abort Pickup Selected MB2[31].21'; 1014 '~S001R13CN.M.RetFmPounceSeld - Robot Return From Pounce Selected MB2[31].22'; 1015 '~S001R13CN.I.StudWld1 Comm Not OK MB2[31].23'; 1016 '~S001R13CN.I.StudWld2 Comm Not OK MB2[31].24'; 1017 '~S001R13CN.I.WldMode - Robot In No Weld MB2[31].25'; 1018 '~S001R13CN.I.PulledTipBypSS - Robot Pulled Tip Bypass Selected MB2[31].26'; 1019 '~S001R13CN.I.FlowNoFlowSS - Robot In No Flow MB2[31].27'; 1020 '~S001R13CN.I.RvtNoRvtSS - Robot In No Rivet MB2[31].28'; 1021 '~S001R13CN.I.WldCtrlCommOk1 - Robot Weld Controller 1 Comm Not OK MB2[31].29'; 1022 '~S001R13CN.I.WldModeStud - Robot In No Weld Stud MB2[31].30'; 1023 '~S001R13CN.Ix.MigWldNoWld - Robot In No Weld Mig MB2[31].31'; 1024 '~S001R13CN.I.StudWld1Rdy - Robot Stud Weld Controller 1 Not Ready MB2[32].0'; 1025 '~S001R13CN.I.Rvt1RdyToOperate - Robot Rivet Controller 1 Not Ready MB2[32].1'; 1026 '~S001R13CN.Ix.MigRdy - Robot Mig Weld Controller Not Ready MB2[32].2'; 1027 '~S001R13CN.Ix.MigWldNoWld - Robot In No Weld MB2[32].3'; 1028 '~Spare MB2[32].4'; 1029 '~S001R13CN.I.WldCtrlCommOk2 - Robot Weld Controller 2 Comm Not OK MB2[32].5'; 